REGION Network 4: Stop 0 - Control logic - Bit profisafe NHE
   RUNG wire#powerrail
      Contact( #tempEStopAllReleased )
      Contact( #tempLcAllFree )
      wire#w1
      Coil( "Tag_5" )
   END_RUNG
   RUNG wire#powerrail
      Contact( #tempLcAccessGrantedZ2 )
   END_RUNG wire#w1
   RUNG wire#powerrail
      Contact( #tempLcAccessGrantedZ3 )
   END_RUNG wire#w1
   // the same network as SCL:
   "Tag_5" := (#tempEStopAllReleased AND #tempLcAllFree) OR #tempLcAccessGrantedZ2 OR #tempLcAccessGrantedZ3;
END_REGION

REGION Network 5
   RUNG wire#powerrail
      #instSafetyDoor(SAF_DOOR_CLSD_RDY =>)
   END_RUNG
   // the same network as SCL:
   #instSafetyDoor();   // "SafetyDoor"
END_REGION

REGION Network 6
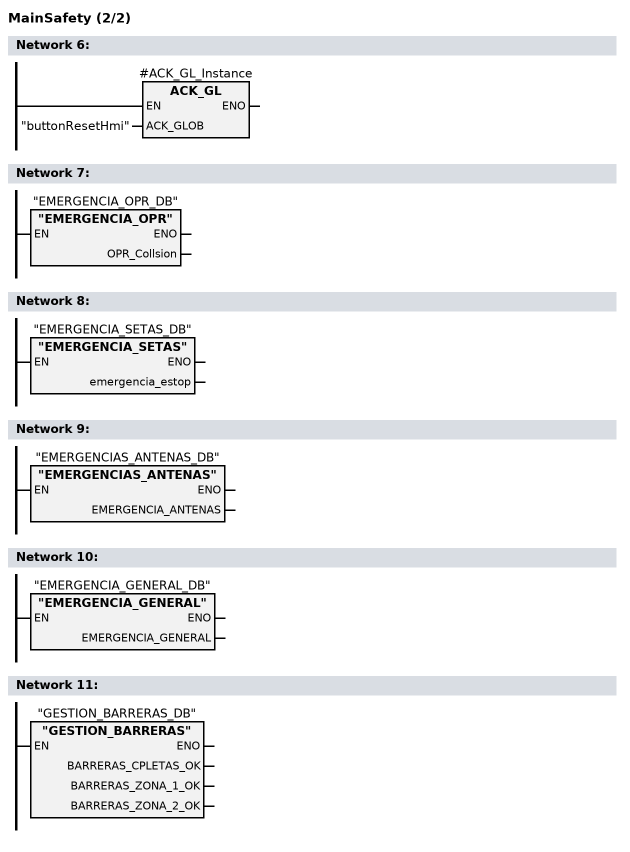
   #ACK_GL_Instance(ACK_GLOB := "buttonResetHmi");   // ACK_GL
END_REGION

REGION Network 7
   RUNG wire#powerrail
      "EMERGENCIA_OPR_DB"(OPR_Collsion =>)
   END_RUNG
   // the same network as SCL:
   "EMERGENCIA_OPR_DB"();   // "EMERGENCIA_OPR"
END_REGION

REGION Network 8
   RUNG wire#powerrail
      "EMERGENCIA_SETAS_DB"(emergencia_estop =>)
   END_RUNG
   // the same network as SCL:
   "EMERGENCIA_SETAS_DB"();   // "EMERGENCIA_SETAS"
END_REGION

REGION Network 9
   RUNG wire#powerrail
      "EMERGENCIAS_ANTENAS_DB"(EMERGENCIA_ANTENAS =>)
   END_RUNG
   // the same network as SCL:
   "EMERGENCIAS_ANTENAS_DB"();   // "EMERGENCIAS_ANTENAS"
END_REGION

REGION Network 10
   RUNG wire#powerrail
      "EMERGENCIA_GENERAL_DB"(EMERGENCIA_GENERAL =>)
   END_RUNG
   // the same network as SCL:
   "EMERGENCIA_GENERAL_DB"();   // "EMERGENCIA_GENERAL"
END_REGION

REGION Network 11
   RUNG wire#powerrail
      "GESTION_BARRERAS_DB"(BARRERAS_CPLETAS_OK =>, BARRERAS_ZONA_1_OK =>, BARRERAS_ZONA_2_OK =>)
   END_RUNG
   // the same network as SCL:
   "GESTION_BARRERAS_DB"();   // "GESTION_BARRERAS"
END_REGION
END_FUNCTION_BLOCK

FUNCTION_BLOCK "SafetyRobot"   // FB3, F_LAD
{ S7_Optimized_Access := 'TRUE' }
VERSION : 0.1
   VAR
      Edge_ACK : Bool;
      mem_ack_trig : Bool;
      ACK_GL_Instance : Bool;
      F_IEC_Timer_Instance_1 : TP;
   END_VAR
   VAR_TEMP   // added for the SCL form of the ladder/FBD networks
      _w1 : Bool;
   END_VAR
BEGIN

REGION Network 1: Reservado (debe ser 1)
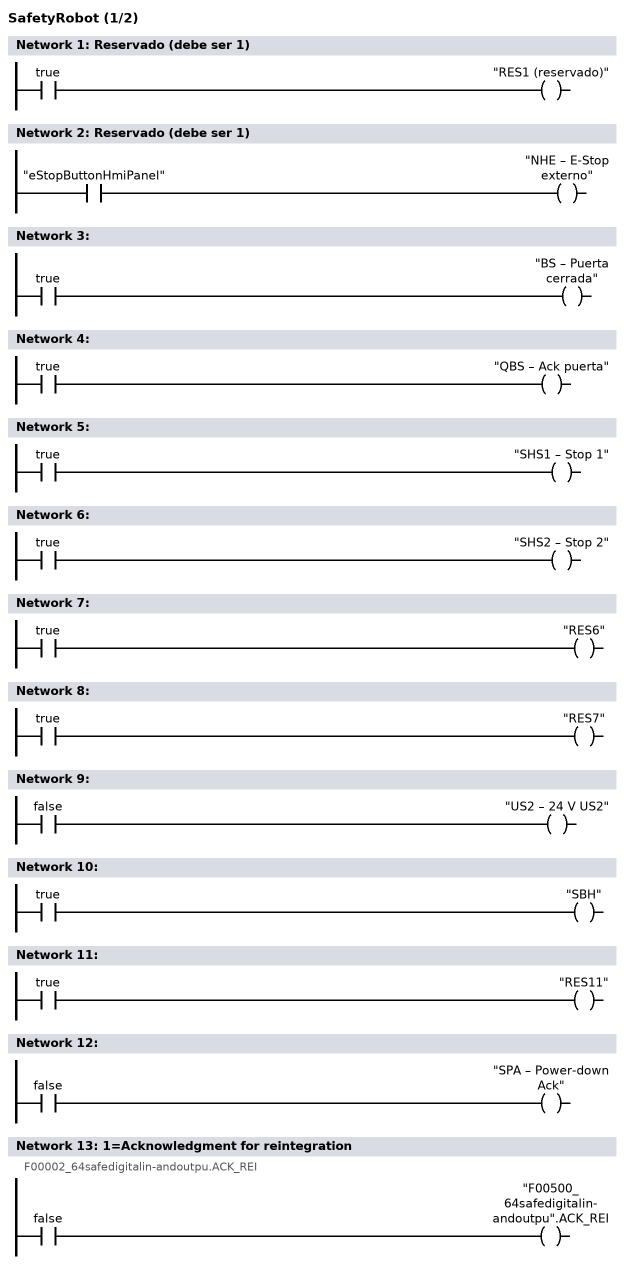
   RUNG wire#powerrail
      Contact( true )
      Coil( "RES1 (reservado)" )
   END_RUNG
   // the same network as SCL:
   "RES1 (reservado)" := true;
END_REGION

REGION Network 2: Reservado (debe ser 1)
   RUNG wire#powerrail
      Contact( "eStopButtonHmiPanel" )
      Coil( "NHE – E‑Stop externo" )
   END_RUNG
   // the same network as SCL:
   "NHE – E‑Stop externo" := "eStopButtonHmiPanel";
END_REGION

REGION Network 3
   RUNG wire#powerrail
      Contact( true )
      Coil( "BS – Puerta cerrada" )
   END_RUNG
   // the same network as SCL:
   "BS – Puerta cerrada" := true;
END_REGION

REGION Network 4
   RUNG wire#powerrail
      Contact( true )
      Coil( "QBS – Ack puerta" )
   END_RUNG
   // the same network as SCL:
   "QBS – Ack puerta" := true;
END_REGION

REGION Network 5
   RUNG wire#powerrail
      Contact( true )
      Coil( "SHS1 – Stop 1" )
   END_RUNG
   // the same network as SCL:
   "SHS1 – Stop 1" := true;
END_REGION

REGION Network 6
   RUNG wire#powerrail
      Contact( true )
      Coil( "SHS2 – Stop 2" )
   END_RUNG
   // the same network as SCL:
   "SHS2 – Stop 2" := true;
END_REGION

REGION Network 7
   RUNG wire#powerrail
      Contact( true )
      Coil( "RES6" )
   END_RUNG
   // the same network as SCL:
   "RES6" := true;
END_REGION

REGION Network 8
   RUNG wire#powerrail
      Contact( true )
      Coil( "RES7" )
   END_RUNG
   // the same network as SCL:
   "RES7" := true;
END_REGION

REGION Network 9
   RUNG wire#powerrail
      Contact( false )
      Coil( "US2 – 24 V US2" )
   END_RUNG
   // the same network as SCL:
   "US2 – 24 V US2" := false;
END_REGION

REGION Network 10
   RUNG wire#powerrail
      Contact( true )
      Coil( "SBH" )
   END_RUNG
   // the same network as SCL:
   "SBH" := true;
END_REGION

REGION Network 11
   RUNG wire#powerrail
      Contact( true )
      Coil( "RES11" )
   END_RUNG
   // the same network as SCL:
   "RES11" := true;
END_REGION

REGION Network 12
   RUNG wire#powerrail
      Contact( false )
      Coil( "SPA – Power‑down Ack" )
   END_RUNG
   // the same network as SCL:
   "SPA – Power‑down Ack" := false;
END_REGION

REGION Network 13: 1=Acknowledgment for reintegration
   // F00002_64safedigitalin-andoutpu.ACK_REI
   RUNG wire#powerrail
      Contact( false )
      Coil( "F00500_64safedigitalin-andoutpu".ACK_REI )
   END_RUNG
   // the same network as SCL:
   "F00500_64safedigitalin-andoutpu".ACK_REI := false;
END_REGION

REGION Network 14: Pulse output
   // - CLK → F00002_…ACK_REQ : Detecta el flanco 0 → 1 que el módulo pone cuando necesita
   // - M → mem_ACK_Trig
   // : reconocimiento. El 1 sólo dura un scan y se guarda internamente en mem_ACK_Trig….
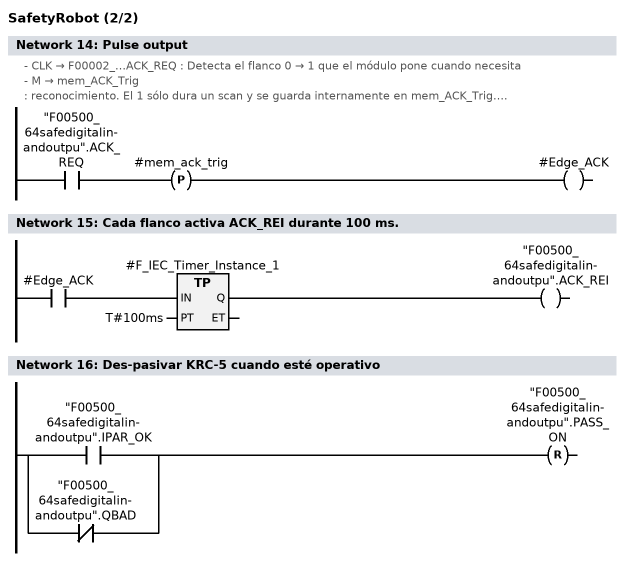
   RUNG wire#powerrail
      Contact( "F00500_64safedigitalin-andoutpu".ACK_REQ )
      P_Trig( #mem_ack_trig )
      Coil( #Edge_ACK )
   END_RUNG
   // the same network as SCL:
   #_w1 := "F00500_64safedigitalin-andoutpu".ACK_REQ AND NOT #mem_ack_trig;   // rising edge
   #mem_ack_trig := "F00500_64safedigitalin-andoutpu".ACK_REQ;
   #Edge_ACK := #_w1;
END_REGION

REGION Network 15: Cada flanco activa ACK_REI durante 100 ms.
   #F_IEC_Timer_Instance_1.TP(IN := #Edge_ACK, PT := T#100ms);
   "F00500_64safedigitalin-andoutpu".ACK_REI := #F_IEC_Timer_Instance_1.Q;
END_REGION

REGION Network 16: Des-pasivar KRC-5 cuando esté operativo
   RUNG wire#powerrail
      Contact( "F00500_64safedigitalin-andoutpu".IPAR_OK )
      wire#w1
      R_Coil( "F00500_64safedigitalin-andoutpu".PASS_ON )
   END_RUNG
   RUNG wire#powerrail
      I_Contact( "F00500_64safedigitalin-andoutpu".QBAD )
   END_RUNG wire#w1
   // the same network as SCL:
   IF "F00500_64safedigitalin-andoutpu".IPAR_OK OR NOT "F00500_64safedigitalin-andoutpu".QBAD THEN
       "F00500_64safedigitalin-andoutpu".PASS_ON := FALSE;
   END_IF;
END_REGION
END_FUNCTION_BLOCK

FUNCTION_BLOCK "EMERGENCIA_SETAS"   // FB16, F_FBD
{ S7_Optimized_Access := 'TRUE' }
VERSION : 0.1
   VAR_OUTPUT
      emergencia_estop : Bool;
   END_VAR
BEGIN

REGION Network 1
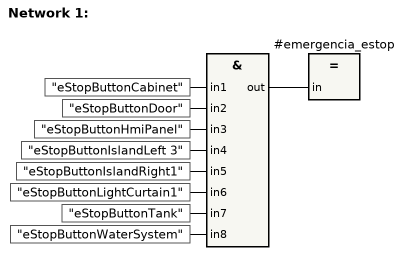
   #emergencia_estop := "eStopButtonCabinet" AND "eStopButtonDoor" AND "eStopButtonHmiPanel" AND "eStopButtonIslandLeft 3" AND "eStopButtonIslandRight1" AND "eStopButtonLightCurtain1" AND "eStopButtonTank" AND "eStopButtonWaterSystem";
END_REGION
END_FUNCTION_BLOCK

FUNCTION_BLOCK "EMERGENCIAS_ANTENAS"   // FB17, F_LAD
{ S7_Optimized_Access := 'TRUE' }
VERSION : 0.1
   VAR_OUTPUT
      EMERGENCIA_ANTENAS : Bool;
   END_VAR
BEGIN

REGION Network 1: YUGO_PUESTO
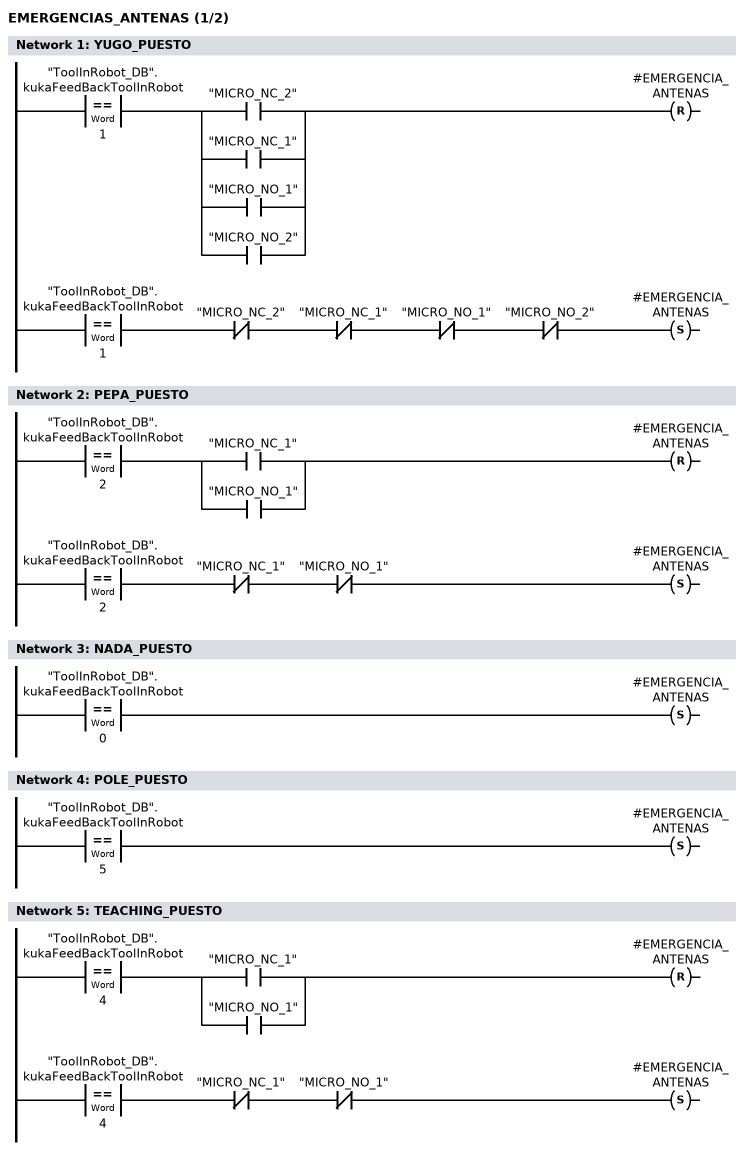
   RUNG wire#powerrail
      { S7_Templates := "SrcType := Word" } EQ_Contact(in1 := "ToolInRobot_DB".kukaFeedBackToolInRobot, in2 := 1)
      wire#w1
      Contact( "MICRO_NC_2" )
      wire#w2
      R_Coil( #EMERGENCIA_ANTENAS )
   END_RUNG
   RUNG wire#w1
      Contact( "MICRO_NC_1" )
   END_RUNG wire#w2
   RUNG wire#w1
      Contact( "MICRO_NO_1" )
   END_RUNG wire#w2
   RUNG wire#w1
      Contact( "MICRO_NO_2" )
   END_RUNG wire#w2
   RUNG wire#powerrail
      { S7_Templates := "SrcType := Word" } EQ_Contact(in1 := "ToolInRobot_DB".kukaFeedBackToolInRobot, in2 := 1)
      I_Contact( "MICRO_NC_2" )
      I_Contact( "MICRO_NC_1" )
      I_Contact( "MICRO_NO_1" )
      I_Contact( "MICRO_NO_2" )
      S_Coil( #EMERGENCIA_ANTENAS )
   END_RUNG
   // the same network as SCL:
   IF ("ToolInRobot_DB".kukaFeedBackToolInRobot = 1) AND ("MICRO_NC_2" OR "MICRO_NC_1" OR "MICRO_NO_1" OR "MICRO_NO_2") THEN
       #EMERGENCIA_ANTENAS := FALSE;
   END_IF;
   IF ("ToolInRobot_DB".kukaFeedBackToolInRobot = 1) AND NOT "MICRO_NC_2" AND NOT "MICRO_NC_1" AND NOT "MICRO_NO_1" AND NOT "MICRO_NO_2" THEN
       #EMERGENCIA_ANTENAS := TRUE;
   END_IF;
END_REGION

REGION Network 2: PEPA_PUESTO
   RUNG wire#powerrail
      { S7_Templates := "SrcType := Word" } EQ_Contact(in1 := "ToolInRobot_DB".kukaFeedBackToolInRobot, in2 := 2)
      wire#w1
      Contact( "MICRO_NC_1" )
      wire#w2
      R_Coil( #EMERGENCIA_ANTENAS )
   END_RUNG
   RUNG wire#w1
      Contact( "MICRO_NO_1" )
   END_RUNG wire#w2
   RUNG wire#powerrail
      { S7_Templates := "SrcType := Word" } EQ_Contact(in1 := "ToolInRobot_DB".kukaFeedBackToolInRobot, in2 := 2)
      I_Contact( "MICRO_NC_1" )
      I_Contact( "MICRO_NO_1" )
      S_Coil( #EMERGENCIA_ANTENAS )
   END_RUNG
   // the same network as SCL:
   IF ("ToolInRobot_DB".kukaFeedBackToolInRobot = 2) AND ("MICRO_NC_1" OR "MICRO_NO_1") THEN
       #EMERGENCIA_ANTENAS := FALSE;
   END_IF;
   IF ("ToolInRobot_DB".kukaFeedBackToolInRobot = 2) AND NOT "MICRO_NC_1" AND NOT "MICRO_NO_1" THEN
       #EMERGENCIA_ANTENAS := TRUE;
   END_IF;
END_REGION

REGION Network 3: NADA_PUESTO
   RUNG wire#powerrail
      { S7_Templates := "SrcType := Word" } EQ_Contact(in1 := "ToolInRobot_DB".kukaFeedBackToolInRobot, in2 := 0)
      S_Coil( #EMERGENCIA_ANTENAS )
   END_RUNG
   // the same network as SCL:
   IF "ToolInRobot_DB".kukaFeedBackToolInRobot = 0 THEN #EMERGENCIA_ANTENAS := TRUE; END_IF;
END_REGION

REGION Network 4: POLE_PUESTO
   RUNG wire#powerrail
      { S7_Templates := "SrcType := Word" } EQ_Contact(in1 := "ToolInRobot_DB".kukaFeedBackToolInRobot, in2 := 5)
      S_Coil( #EMERGENCIA_ANTENAS )
   END_RUNG
   // the same network as SCL:
   IF "ToolInRobot_DB".kukaFeedBackToolInRobot = 5 THEN #EMERGENCIA_ANTENAS := TRUE; END_IF;
END_REGION

REGION Network 5: TEACHING_PUESTO
   RUNG wire#powerrail
      { S7_Templates := "SrcType := Word" } EQ_Contact(in1 := "ToolInRobot_DB".kukaFeedBackToolInRobot, in2 := 4)
      wire#w1
      Contact( "MICRO_NC_1" )
      wire#w2
      R_Coil( #EMERGENCIA_ANTENAS )
   END_RUNG
   RUNG wire#w1
      Contact( "MICRO_NO_1" )
   END_RUNG wire#w2
   RUNG wire#powerrail
      { S7_Templates := "SrcType := Word" } EQ_Contact(in1 := "ToolInRobot_DB".kukaFeedBackToolInRobot, in2 := 4)
      I_Contact( "MICRO_NC_1" )
      I_Contact( "MICRO_NO_1" )
      S_Coil( #EMERGENCIA_ANTENAS )
   END_RUNG
   // the same network as SCL:
   IF ("ToolInRobot_DB".kukaFeedBackToolInRobot = 4) AND ("MICRO_NC_1" OR "MICRO_NO_1") THEN
       #EMERGENCIA_ANTENAS := FALSE;
   END_IF;
   IF ("ToolInRobot_DB".kukaFeedBackToolInRobot = 4) AND NOT "MICRO_NC_1" AND NOT "MICRO_NO_1" THEN
       #EMERGENCIA_ANTENAS := TRUE;
   END_IF;
END_REGION

REGION Network 6: MARKER_PUESTO
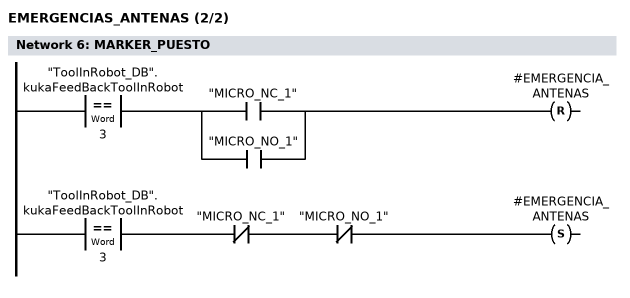
   RUNG wire#powerrail
      { S7_Templates := "SrcType := Word" } EQ_Contact(in1 := "ToolInRobot_DB".kukaFeedBackToolInRobot, in2 := 3)
      wire#w1
      Contact( "MICRO_NC_1" )
      wire#w2
      R_Coil( #EMERGENCIA_ANTENAS )
   END_RUNG
   RUNG wire#w1
      Contact( "MICRO_NO_1" )
   END_RUNG wire#w2
   RUNG wire#powerrail
      { S7_Templates := "SrcType := Word" } EQ_Contact(in1 := "ToolInRobot_DB".kukaFeedBackToolInRobot, in2 := 3)
      I_Contact( "MICRO_NC_1" )
      I_Contact( "MICRO_NO_1" )
      S_Coil( #EMERGENCIA_ANTENAS )
   END_RUNG
   // the same network as SCL:
   IF ("ToolInRobot_DB".kukaFeedBackToolInRobot = 3) AND ("MICRO_NC_1" OR "MICRO_NO_1") THEN
       #EMERGENCIA_ANTENAS := FALSE;
   END_IF;
   IF ("ToolInRobot_DB".kukaFeedBackToolInRobot = 3) AND NOT "MICRO_NC_1" AND NOT "MICRO_NO_1" THEN
       #EMERGENCIA_ANTENAS := TRUE;
   END_IF;
END_REGION
END_FUNCTION_BLOCK

FUNCTION_BLOCK "EMERGENCIA_OPR"   // FB18, F_LAD
{ S7_Optimized_Access := 'TRUE' }
VERSION : 0.1
   VAR_OUTPUT
      OPR_Collsion : Bool;
   END_VAR
BEGIN

REGION Network 1
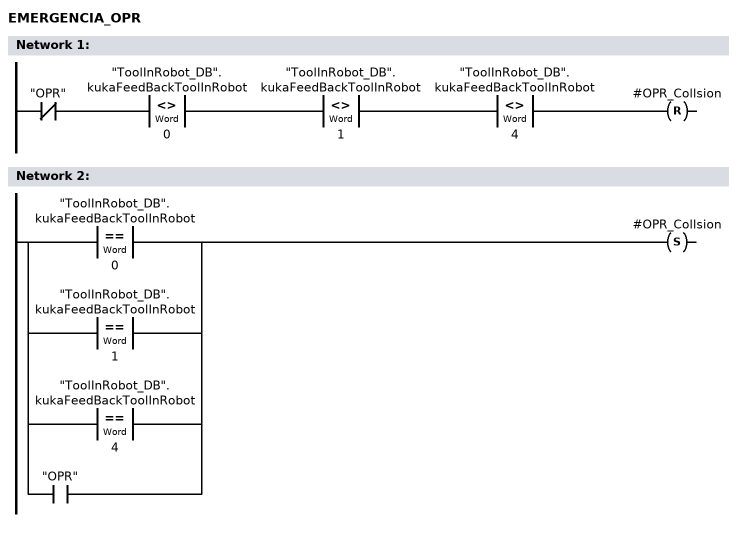
   RUNG wire#powerrail
      I_Contact( "OPR" )
      { S7_Templates := "SrcType := Word" } NE_Contact(in1 := "ToolInRobot_DB".kukaFeedBackToolInRobot, in2 := 0)
      { S7_Templates := "SrcType := Word" } NE_Contact(in1 := "ToolInRobot_DB".kukaFeedBackToolInRobot, in2 := 1)
      { S7_Templates := "SrcType := Word" } NE_Contact(in1 := "ToolInRobot_DB".kukaFeedBackToolInRobot, in2 := 4)
      R_Coil( #OPR_Collsion )
   END_RUNG
   // the same network as SCL:
   IF NOT "OPR" AND ("ToolInRobot_DB".kukaFeedBackToolInRobot <> 0) AND ("ToolInRobot_DB".kukaFeedBackToolInRobot <> 1) AND ("ToolInRobot_DB".kukaFeedBackToolInRobot <> 4) THEN
       #OPR_Collsion := FALSE;
   END_IF;
END_REGION

REGION Network 2
   RUNG wire#powerrail
      { S7_Templates := "SrcType := Word" } EQ_Contact(in1 := "ToolInRobot_DB".kukaFeedBackToolInRobot, in2 := 0)
      wire#w1
      S_Coil( #OPR_Collsion )
   END_RUNG
   RUNG wire#powerrail
      { S7_Templates := "SrcType := Word" } EQ_Contact(in1 := "ToolInRobot_DB".kukaFeedBackToolInRobot, in2 := 1)
   END_RUNG wire#w1
   RUNG wire#powerrail
      { S7_Templates := "SrcType := Word" } EQ_Contact(in1 := "ToolInRobot_DB".kukaFeedBackToolInRobot, in2 := 4)
   END_RUNG wire#w1
   RUNG wire#powerrail
      Contact( "OPR" )
   END_RUNG wire#w1
   // the same network as SCL:
   IF ("ToolInRobot_DB".kukaFeedBackToolInRobot = 0) OR ("ToolInRobot_DB".kukaFeedBackToolInRobot = 1) OR ("ToolInRobot_DB".kukaFeedBackToolInRobot = 4) OR "OPR" THEN
       #OPR_Collsion := TRUE;
   END_IF;
END_REGION
END_FUNCTION_BLOCK

FUNCTION_BLOCK "ACCESO_ZONA_1"   // FB19, F_FBD
{ S7_Optimized_Access := 'TRUE' }
VERSION : 0.1
BEGIN
END_FUNCTION_BLOCK

FUNCTION_BLOCK "ACCESO_ZONA_2"   // FB23, F_LAD
{ S7_Optimized_Access := 'TRUE' }
VERSION : 0.1
BEGIN
END_FUNCTION_BLOCK

FUNCTION_BLOCK "ACCESO_COMPLETO"   // FB24, F_FBD
{ S7_Optimized_Access := 'TRUE' }
VERSION : 0.1
   VAR_OUTPUT
      ACCESO_PERMITIDO : Bool;
   END_VAR
BEGIN

REGION Network 1
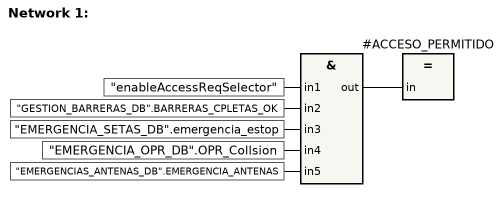
   #ACCESO_PERMITIDO := "enableAccessReqSelector" AND "GESTION_BARRERAS_DB".BARRERAS_CPLETAS_OK AND "EMERGENCIA_SETAS_DB".emergencia_estop AND "EMERGENCIA_OPR_DB".OPR_Collsion AND "EMERGENCIAS_ANTENAS_DB".EMERGENCIA_ANTENAS;
END_REGION
END_FUNCTION_BLOCK

FUNCTION_BLOCK "GESTION_BARRERAS"   // FB25, F_FBD
{ S7_Optimized_Access := 'TRUE' }
VERSION : 0.1
   VAR_OUTPUT
      BARRERAS_CPLETAS_OK : Bool;
      BARRERAS_ZONA_1_OK : Bool;
      BARRERAS_ZONA_2_OK : Bool;
   END_VAR
BEGIN

REGION Network 1
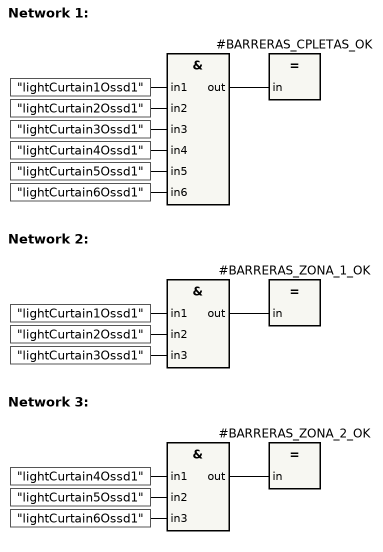
   #BARRERAS_CPLETAS_OK := "lightCurtain1Ossd1" AND "lightCurtain2Ossd1" AND "lightCurtain3Ossd1" AND "lightCurtain4Ossd1" AND "lightCurtain5Ossd1" AND "lightCurtain6Ossd1";
END_REGION

REGION Network 2
   #BARRERAS_ZONA_1_OK := "lightCurtain1Ossd1" AND "lightCurtain2Ossd1" AND "lightCurtain3Ossd1";
END_REGION

REGION Network 3
   #BARRERAS_ZONA_2_OK := "lightCurtain4Ossd1" AND "lightCurtain5Ossd1" AND "lightCurtain6Ossd1";
END_REGION
END_FUNCTION_BLOCK

FUNCTION_BLOCK "EMERGENCIA_GENERAL"   // FB26, F_FBD
{ S7_Optimized_Access := 'TRUE' }
VERSION : 0.1
   VAR_OUTPUT
      EMERGENCIA_GENERAL : Bool;
   END_VAR
BEGIN

REGION Network 1
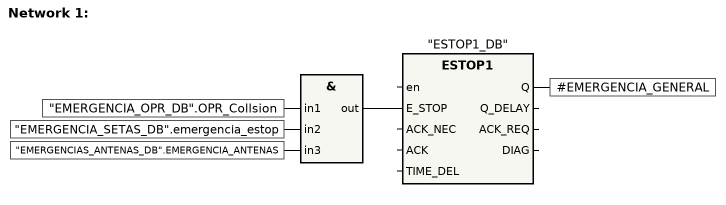
   "ESTOP1_DB"(E_STOP := "EMERGENCIA_OPR_DB".OPR_Collsion AND "EMERGENCIA_SETAS_DB".emergencia_estop AND "EMERGENCIAS_ANTENAS_DB".EMERGENCIA_ANTENAS,   // ESTOP1
               Q => #EMERGENCIA_GENERAL);
END_REGION
END_FUNCTION_BLOCK

FUNCTION_BLOCK "REARMAR_MAQUINA"   // FB27, F_FBD
{ S7_Optimized_Access := 'TRUE' }
VERSION : 0.1
BEGIN
END_FUNCTION_BLOCK

FUNCTION_BLOCK "EMERGENCIAS_ROBOT"   // FB29, F_LAD
{ S7_Optimized_Access := 'TRUE' }
VERSION : 0.1
BEGIN

REGION Network 1: Reservado (debe ser 1)
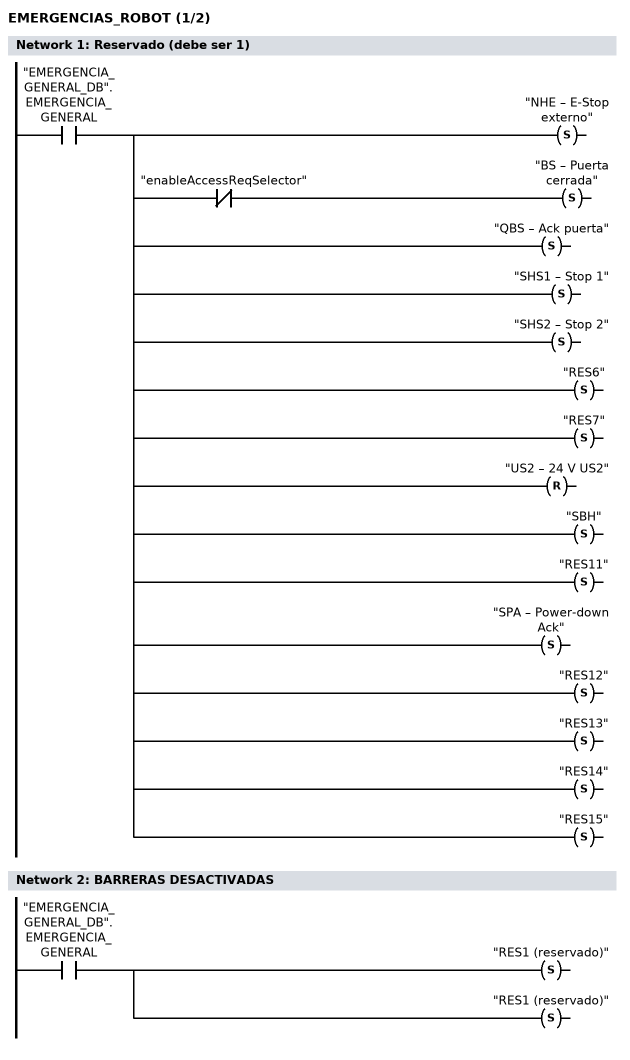
   RUNG wire#powerrail
      Contact( "EMERGENCIA_GENERAL_DB".EMERGENCIA_GENERAL )
      wire#w1
      S_Coil( "NHE – E‑Stop externo" )
   END_RUNG
   RUNG wire#w1
      I_Contact( "enableAccessReqSelector" )
      S_Coil( "BS – Puerta cerrada" )
   END_RUNG
   RUNG wire#w1
      S_Coil( "QBS – Ack puerta" )
   END_RUNG
   RUNG wire#w1
      S_Coil( "SHS1 – Stop 1" )
   END_RUNG
   RUNG wire#w1
      S_Coil( "SHS2 – Stop 2" )
   END_RUNG
   RUNG wire#w1
      S_Coil( "RES6" )
   END_RUNG
   RUNG wire#w1
      S_Coil( "RES7" )
   END_RUNG
   RUNG wire#w1
      R_Coil( "US2 – 24 V US2" )
   END_RUNG
   RUNG wire#w1
      S_Coil( "SBH" )
   END_RUNG
   RUNG wire#w1
      S_Coil( "RES11" )
   END_RUNG
   RUNG wire#w1
      S_Coil( "SPA – Power‑down Ack" )
   END_RUNG
   RUNG wire#w1
      S_Coil( "RES12" )
   END_RUNG
   RUNG wire#w1
      S_Coil( "RES13" )
   END_RUNG
   RUNG wire#w1
      S_Coil( "RES14" )
   END_RUNG
   RUNG wire#w1
      S_Coil( "RES15" )
   END_RUNG
   // the same network as SCL:
   IF "EMERGENCIA_GENERAL_DB".EMERGENCIA_GENERAL THEN "NHE – E‑Stop externo" := TRUE; END_IF;
   IF "EMERGENCIA_GENERAL_DB".EMERGENCIA_GENERAL AND NOT "enableAccessReqSelector" THEN
       "BS – Puerta cerrada" := TRUE;
   END_IF;
   IF "EMERGENCIA_GENERAL_DB".EMERGENCIA_GENERAL THEN
       "QBS – Ack puerta" := TRUE;
       "SHS1 – Stop 1" := TRUE;
       "SHS2 – Stop 2" := TRUE;
       "RES6" := TRUE;
       "RES7" := TRUE;
       "US2 – 24 V US2" := FALSE;
       "SBH" := TRUE;
       "RES11" := TRUE;
       "SPA – Power‑down Ack" := TRUE;
       "RES12" := TRUE;
       "RES13" := TRUE;
       "RES14" := TRUE;
       "RES15" := TRUE;
   END_IF;
END_REGION

REGION Network 2: BARRERAS DESACTIVADAS
   RUNG wire#powerrail
      Contact( "EMERGENCIA_GENERAL_DB".EMERGENCIA_GENERAL )
      wire#w1
      S_Coil( "RES1 (reservado)" )
   END_RUNG
   RUNG wire#w1
      S_Coil( "RES1 (reservado)" )
   END_RUNG
   // the same network as SCL:
   IF "EMERGENCIA_GENERAL_DB".EMERGENCIA_GENERAL THEN
       "RES1 (reservado)" := TRUE;
       "RES1 (reservado)" := TRUE;
   END_IF;
END_REGION

REGION Network 4: Reservado (debe ser 1)
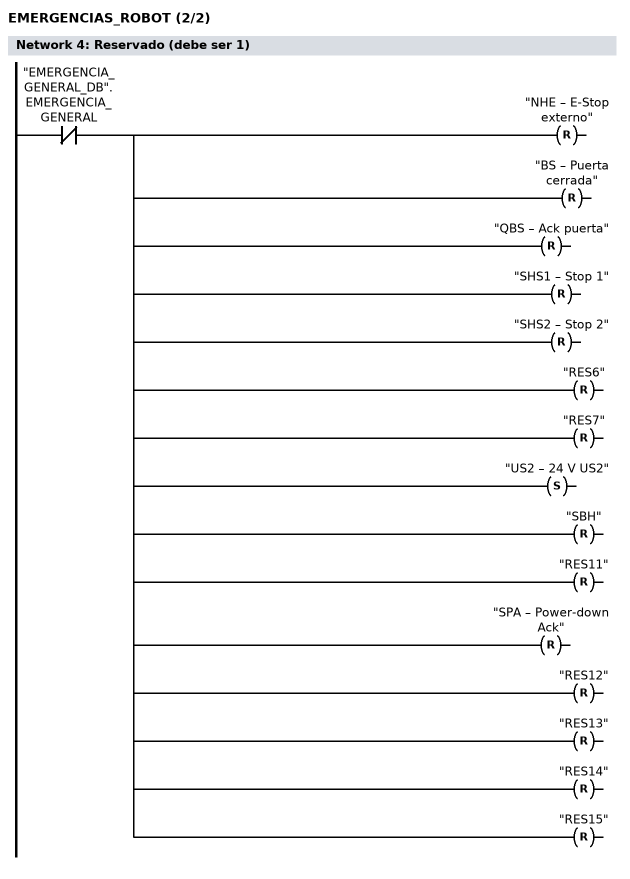
   RUNG wire#powerrail
      I_Contact( "EMERGENCIA_GENERAL_DB".EMERGENCIA_GENERAL )
      wire#w1
      R_Coil( "NHE – E‑Stop externo" )
   END_RUNG
   RUNG wire#w1
      R_Coil( "BS – Puerta cerrada" )
   END_RUNG
   RUNG wire#w1
      R_Coil( "QBS – Ack puerta" )
   END_RUNG
   RUNG wire#w1
      R_Coil( "SHS1 – Stop 1" )
   END_RUNG
   RUNG wire#w1
      R_Coil( "SHS2 – Stop 2" )
   END_RUNG
   RUNG wire#w1
      R_Coil( "RES6" )
   END_RUNG
   RUNG wire#w1
      R_Coil( "RES7" )
   END_RUNG
   RUNG wire#w1
      S_Coil( "US2 – 24 V US2" )
   END_RUNG
   RUNG wire#w1
      R_Coil( "SBH" )
   END_RUNG
   RUNG wire#w1
      R_Coil( "RES11" )
   END_RUNG
   RUNG wire#w1
      R_Coil( "SPA – Power‑down Ack" )
   END_RUNG
   RUNG wire#w1
      R_Coil( "RES12" )
   END_RUNG
   RUNG wire#w1
      R_Coil( "RES13" )
   END_RUNG
   RUNG wire#w1
      R_Coil( "RES14" )
   END_RUNG
   RUNG wire#w1
      R_Coil( "RES15" )
   END_RUNG
   // the same network as SCL:
   IF NOT "EMERGENCIA_GENERAL_DB".EMERGENCIA_GENERAL THEN
       "NHE – E‑Stop externo" := FALSE;
       "BS – Puerta cerrada" := FALSE;
       "QBS – Ack puerta" := FALSE;
       "SHS1 – Stop 1" := FALSE;
       "SHS2 – Stop 2" := FALSE;
       "RES6" := FALSE;
       "RES7" := FALSE;
       "US2 – 24 V US2" := TRUE;
       "SBH" := FALSE;
       "RES11" := FALSE;
       "SPA – Power‑down Ack" := FALSE;
       "RES12" := FALSE;
       "RES13" := FALSE;
       "RES14" := FALSE;
       "RES15" := FALSE;
   END_IF;
END_REGION
END_FUNCTION_BLOCK

// folder: 30. Safety/SafetyFunctions

FUNCTION_BLOCK "EStopGroup"   // FB2, F_LAD
{ S7_Optimized_Access := 'TRUE' }
VERSION : 0.1
   VAR_INPUT
      acknowledge : Bool;   // Acknowledge / Quittierung, Positive Flanke notwendig, NO / Acknowledge, positive signal edge, NO
      eStop1 : Bool;   // eStop / Not-Halt Drucktaster, False: Not-Halt ausgelöst NC / eStop input, False: eStop triggered NC
      eStop2 : Bool;   // eStop / Not-Halt Drucktaster, False: Not-Halt ausgelöst NC / eStop input, False: eStop triggered NC
      eStop3 : Bool;   // eStop / Not-Halt Drucktaster, False: Not-Halt ausgelöst NC / eStop input, False: eStop triggered NC
      eStop4 : Bool;   // eStop / Not-Halt Drucktaster, False: Not-Halt ausgelöst NC / eStop input, False: eStop triggered NC
      eStop5 : Bool;   // eStop / Not-Halt Drucktaster, False: Not-Halt ausgelöst NC / eStop input, False: eStop triggered NC
      eStop6 : Bool;   // eStop / Not-Halt Drucktaster, False: Not-Halt ausgelöst NC / eStop input, False: eStop triggered NC
      eStop7 : Bool;   // eStop / Not-Halt Drucktaster, False: Not-Halt ausgelöst NC / eStop input, False: eStop triggered NC
      eStop8 : Bool;   // eStop / Not-Halt Drucktaster, False: Not-Halt ausgelöst NC / eStop input, False: eStop triggered NC
   END_VAR
   VAR_OUTPUT
      eStopAllReleased : Bool;   // Output K1/K2 / Aktor Ausgang an F-DQ / actuator output F-DQ
      eStop1Released : Bool;   // releaseEStop / Freigabe Not-Halt, True: Not-Halt ist entriegelt und quittiert / Release eStop; True: button is released and acknowledged
      eStop2Released : Bool;   // releaseEStop / Freigabe Not-Halt, True: Not-Halt ist entriegelt und quittiert / Release eStop; True: button is released and acknowledged
      eStop3Released : Bool;   // releaseEStop / Freigabe Not-Halt, True: Not-Halt ist entriegelt und quittiert / Release eStop; True: button is released and acknowledged
      eStop4Released : Bool;
      eStop5Released : Bool;
      eStop6Released : Bool;
      eStop7Released : Bool;
      eStop8Released : Bool;
      acknowledgeReqestedEStop : Bool;   // eStop acknowlege requested / Quittierung Not-Halt notwendig, True: Quittierung notwendig / eStop button acknowlege requested; True: acknowledge requested
   END_VAR
   VAR
      statReleaseEStop1 : Bool;   // Static value for eStop status / Interne Variable für den Status des Not-Halt
      statReleaseEStop2 : Bool;   // Static value for eStop status / Interne Variable für den Status des Not-Halt
      statReleaseEStop3 : Bool;   // Static value for eStop status / Interne Variable für den Status des Not-Halt
      statReleaseEStop4 : Bool;   // Static value for eStop status / Interne Variable für den Status des Not-Halt
      statReleaseEStop5 : Bool;   // Static value for eStop status / Interne Variable für den Status des Not-Halt
      statReleaseEStop6 : Bool;   // Static value for eStop status / Interne Variable für den Status des Not-Halt
      statReleaseEStop7 : Bool;   // Static value for eStop status / Interne Variable für den Status des Not-Halt
      statReleaseEStop8 : Bool;   // Static value for eStop status / Interne Variable für den Status des Not-Halt
      statAcknowledgeReqestedEStop1 : Bool;   // Static value for eStop acknowlege requested / Interne Variable für die Quittieranforderung des Not-Halt
      statAcknowledgeReqestedEStop2 : Bool;   // Static value for eStop acknowlege requested / Interne Variable für die Quittieranforderung des Not-Halt
      statAcknowledgeReqestedEStop3 : Bool;   // Static value for eStop acknowlege requested / Interne Variable für die Quittieranforderung des Not-Halt
      statAcknowledgeReqestedEStop4 : Bool;   // Static value for eStop acknowlege requested / Interne Variable für die Quittieranforderung des Not-Halt
      statAcknowledgeReqestedEStop5 : Bool;   // Static value for eStop acknowlege requested / Interne Variable für die Quittieranforderung des Not-Halt
      statAcknowledgeReqestedEStop6 : Bool;   // Static value for eStop acknowlege requested / Interne Variable für die Quittieranforderung des Not-Halt
      statAcknowledgeReqestedEStop7 : Bool;
      statAcknowledgeReqestedEStop8 : Bool;
      ESTOP1_Instance_1 : ESTOP1;
      ESTOP1_Instance_2 : ESTOP1;
      ESTOP1_Instance_3 : ESTOP1;
      ESTOP1_Instance_4 : ESTOP1;
      ESTOP1_Instance_5 : ESTOP1;
      ESTOP1_Instance_6 : ESTOP1;
      ESTOP1_Instance_7 : ESTOP1;
      ESTOP1_Instance_8 : ESTOP1;
   END_VAR
BEGIN

REGION Network 1
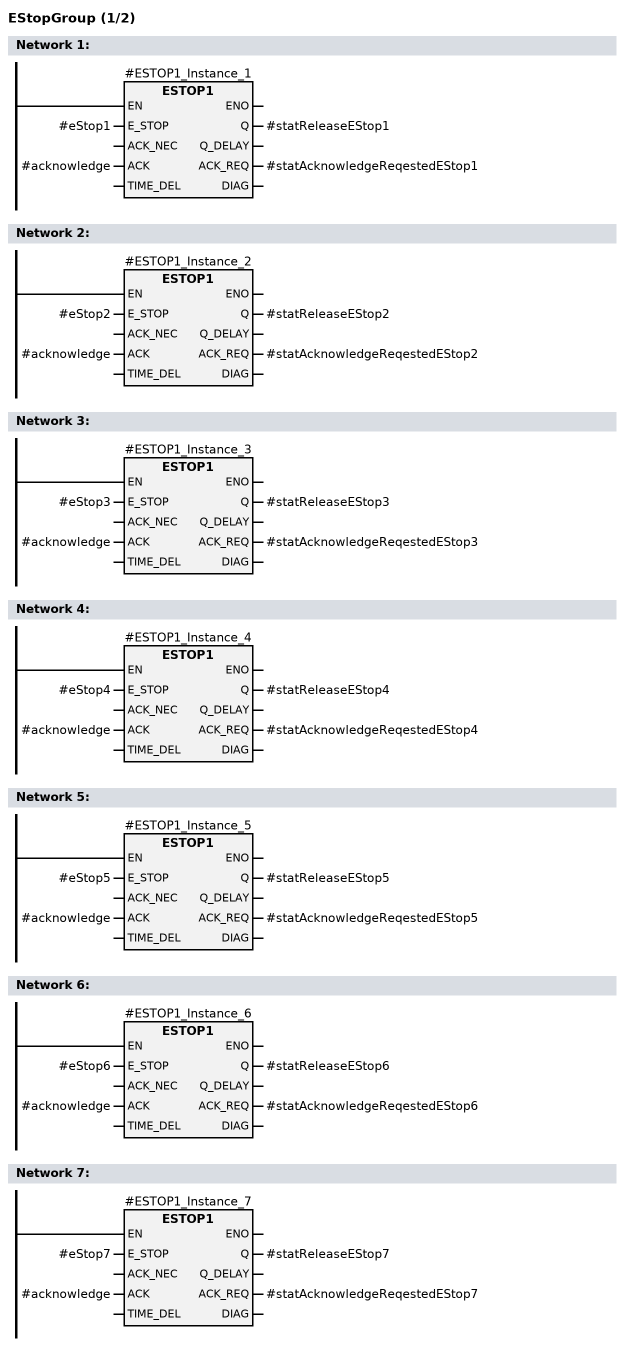
   #ESTOP1_Instance_1(E_STOP := #eStop1,   // ESTOP1
                      ACK := #acknowledge,
                      Q => #statReleaseEStop1,
                      ACK_REQ => #statAcknowledgeReqestedEStop1);
END_REGION

REGION Network 2
   #ESTOP1_Instance_2(E_STOP := #eStop2,   // ESTOP1
                      ACK := #acknowledge,
                      Q => #statReleaseEStop2,
                      ACK_REQ => #statAcknowledgeReqestedEStop2);
END_REGION

REGION Network 3
   #ESTOP1_Instance_3(E_STOP := #eStop3,   // ESTOP1
                      ACK := #acknowledge,
                      Q => #statReleaseEStop3,
                      ACK_REQ => #statAcknowledgeReqestedEStop3);
END_REGION

REGION Network 4
   #ESTOP1_Instance_4(E_STOP := #eStop4,   // ESTOP1
                      ACK := #acknowledge,
                      Q => #statReleaseEStop4,
                      ACK_REQ => #statAcknowledgeReqestedEStop4);
END_REGION

REGION Network 5
   #ESTOP1_Instance_5(E_STOP := #eStop5,   // ESTOP1
                      ACK := #acknowledge,
                      Q => #statReleaseEStop5,
                      ACK_REQ => #statAcknowledgeReqestedEStop5);
END_REGION

REGION Network 6
   #ESTOP1_Instance_6(E_STOP := #eStop6,   // ESTOP1
                      ACK := #acknowledge,
                      Q => #statReleaseEStop6,
                      ACK_REQ => #statAcknowledgeReqestedEStop6);
END_REGION

REGION Network 7
   #ESTOP1_Instance_7(E_STOP := #eStop7,   // ESTOP1
                      ACK := #acknowledge,
                      Q => #statReleaseEStop7,
                      ACK_REQ => #statAcknowledgeReqestedEStop7);
END_REGION

REGION Network 8